// TIA Portal project "SSA-3GHz_V18" (V18) (continued)
REGION Network 10: PS_OK
   RUNG wire#powerrail
      Contact( "DigitalInputs".PS_OK.DigitalIN.NegLogic )
      I_Contact( "DigitalInputs".PS_OK.DigitalIN.PhysIn )
      wire#w1
      Coil( "DigitalInputs".PS_OK.DigitalIN.Out )
   END_RUNG
   RUNG wire#powerrail
      I_Contact( "DigitalInputs".PS_OK.DigitalIN.NegLogic )
      Contact( "DigitalInputs".PS_OK.DigitalIN.PhysIn )
   END_RUNG wire#w1
   // the same network as SCL:
   "DigitalInputs".PS_OK.DigitalIN.Out := ("DigitalInputs".PS_OK.DigitalIN.NegLogic AND NOT "DigitalInputs".PS_OK.DigitalIN.PhysIn) OR (NOT "DigitalInputs".PS_OK.DigitalIN.NegLogic AND "DigitalInputs".PS_OK.DigitalIN.PhysIn);
END_REGION

REGION Network 11: CoolingWtrOK
   RUNG wire#powerrail
      Contact( "CoolingWtrOK" )
      Coil( "DigitalInputs".CoolingWtrOK.DigitalIN.PhysIn )
   END_RUNG
   // the same network as SCL:
   "DigitalInputs".CoolingWtrOK.DigitalIN.PhysIn := "CoolingWtrOK";
END_REGION

REGION Network 12: CoolingWtrOK
   RUNG wire#powerrail
      Contact( "DigitalInputs".CoolingWtrOK.DigitalIN.NegLogic )
      I_Contact( "DigitalInputs".CoolingWtrOK.DigitalIN.PhysIn )
      wire#w1
      Coil( "DigitalInputs".CoolingWtrOK.DigitalIN.Out )
   END_RUNG
   RUNG wire#powerrail
      I_Contact( "DigitalInputs".CoolingWtrOK.DigitalIN.NegLogic )
      Contact( "DigitalInputs".CoolingWtrOK.DigitalIN.PhysIn )
   END_RUNG wire#w1
   // the same network as SCL:
   "DigitalInputs".CoolingWtrOK.DigitalIN.Out := ("DigitalInputs".CoolingWtrOK.DigitalIN.NegLogic AND NOT "DigitalInputs".CoolingWtrOK.DigitalIN.PhysIn) OR (NOT "DigitalInputs".CoolingWtrOK.DigitalIN.NegLogic AND "DigitalInputs".CoolingWtrOK.DigitalIN.PhysIn);
END_REGION

REGION Network 13: FanOK
   RUNG wire#powerrail
      Contact( "FanOK" )
      Coil( "DigitalInputs".FanOK.DigitalIN.PhysIn )
   END_RUNG
   // the same network as SCL:
   "DigitalInputs".FanOK.DigitalIN.PhysIn := "FanOK";
END_REGION

REGION Network 14: FanOK
   RUNG wire#powerrail
      Contact( "DigitalInputs".FanOK.DigitalIN.NegLogic )
      I_Contact( "DigitalInputs".FanOK.DigitalIN.PhysIn )
      wire#w1
      Coil( "DigitalInputs".FanOK.DigitalIN.Out )
   END_RUNG
   RUNG wire#powerrail
      I_Contact( "DigitalInputs".FanOK.DigitalIN.NegLogic )
      Contact( "DigitalInputs".FanOK.DigitalIN.PhysIn )
   END_RUNG wire#w1
   // the same network as SCL:
   "DigitalInputs".FanOK.DigitalIN.Out := ("DigitalInputs".FanOK.DigitalIN.NegLogic AND NOT "DigitalInputs".FanOK.DigitalIN.PhysIn) OR (NOT "DigitalInputs".FanOK.DigitalIN.NegLogic AND "DigitalInputs".FanOK.DigitalIN.PhysIn);
END_REGION

REGION Network 15: ExtIntlkOK
   RUNG wire#powerrail
      Contact( "ExtIntlkOK" )
      Coil( "DigitalInputs".ExtIntlkOK.DigitalIN.PhysIn )
   END_RUNG
   // the same network as SCL:
   "DigitalInputs".ExtIntlkOK.DigitalIN.PhysIn := "ExtIntlkOK";
END_REGION

REGION Network 16: ExtIntlkOK
   RUNG wire#powerrail
      Contact( "DigitalInputs".ExtIntlkOK.DigitalIN.NegLogic )
      I_Contact( "DigitalInputs".ExtIntlkOK.DigitalIN.PhysIn )
      wire#w1
      Coil( "DigitalInputs".ExtIntlkOK.DigitalIN.Out )
   END_RUNG
   RUNG wire#powerrail
      I_Contact( "DigitalInputs".ExtIntlkOK.DigitalIN.NegLogic )
      Contact( "DigitalInputs".ExtIntlkOK.DigitalIN.PhysIn )
   END_RUNG wire#w1
   // the same network as SCL:
   "DigitalInputs".ExtIntlkOK.DigitalIN.Out := ("DigitalInputs".ExtIntlkOK.DigitalIN.NegLogic AND NOT "DigitalInputs".ExtIntlkOK.DigitalIN.PhysIn) OR (NOT "DigitalInputs".ExtIntlkOK.DigitalIN.NegLogic AND "DigitalInputs".ExtIntlkOK.DigitalIN.PhysIn);
END_REGION
END_FUNCTION

FUNCTION "ProcessAI" : Void   // FC401, LAD
{ S7_Optimized_Access := 'TRUE' }
VERSION : 0.1
   VAR_TEMP
      tmpR : Real;
   END_VAR
BEGIN

REGION Network 1: U drain_RBK
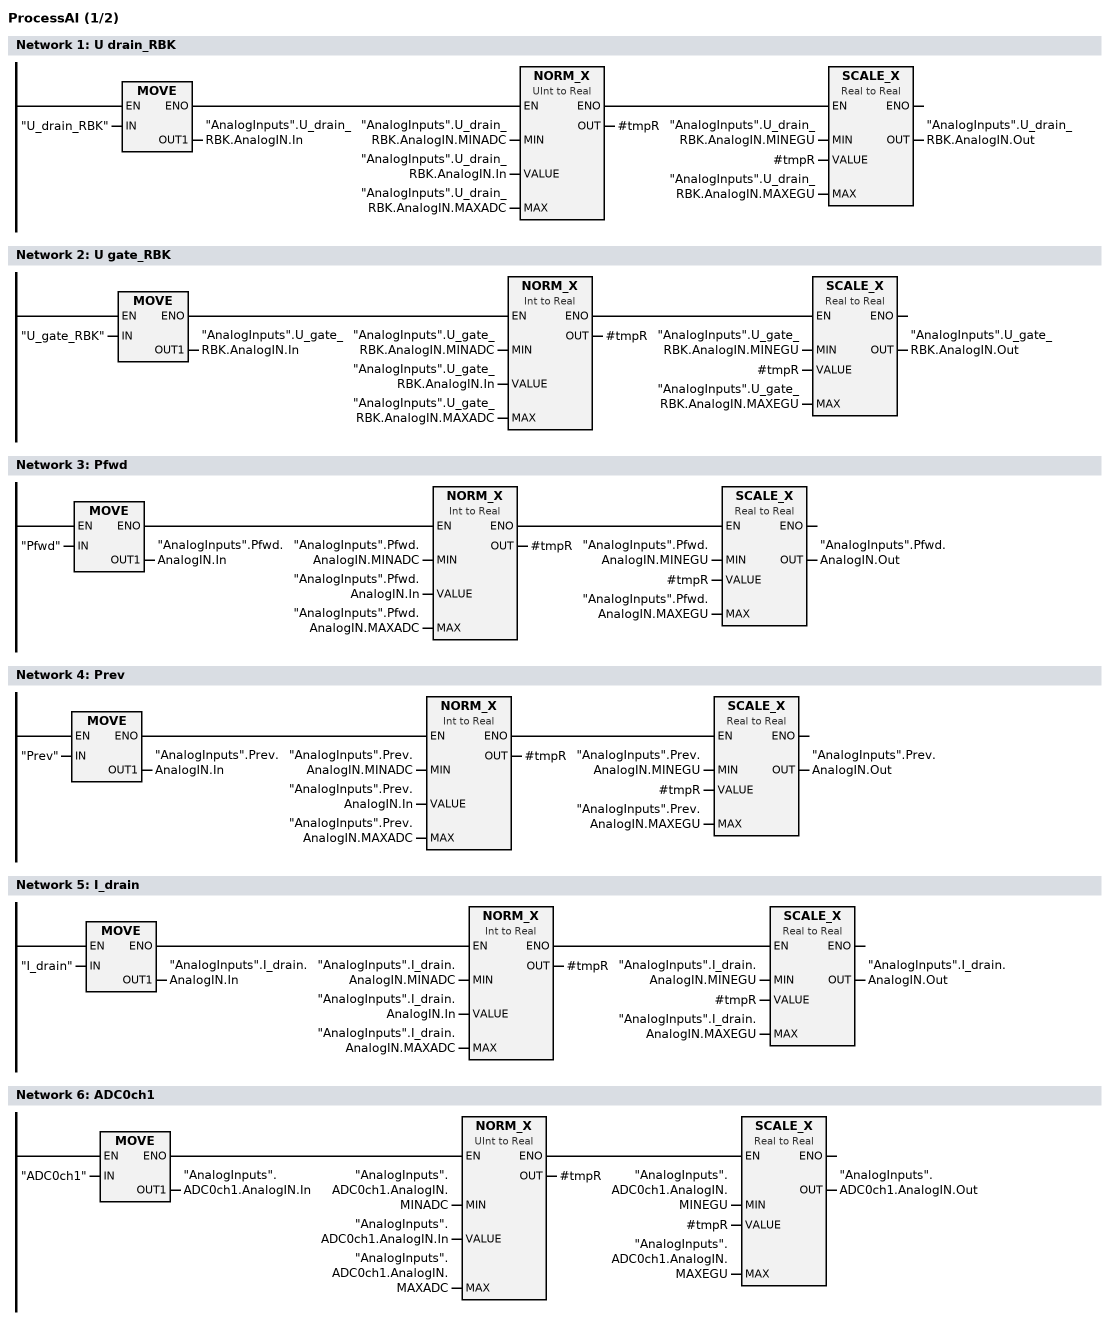
   RUNG wire#powerrail
      Move(in := "U_drain_RBK", out1 => "AnalogInputs".U_drain_RBK.AnalogIN.In)
      { S7_Templates := "[SrcType := UInt, DestType := Real]" } Normalize(min := "AnalogInputs".U_drain_RBK.AnalogIN.MINADC, value := "AnalogInputs".U_drain_RBK.AnalogIN.In, max := "AnalogInputs".U_drain_RBK.AnalogIN.MAXADC, out => #tmpR)
      { S7_Templates := "[SrcType := Real, DestType := Real]" } Scale(min := "AnalogInputs".U_drain_RBK.AnalogIN.MINEGU, value := #tmpR, max := "AnalogInputs".U_drain_RBK.AnalogIN.MAXEGU, out => "AnalogInputs".U_drain_RBK.AnalogIN.Out)
   END_RUNG
   // the same network as SCL:
   "AnalogInputs".U_drain_RBK.AnalogIN.In := "U_drain_RBK";
   #tmpR := NORM_X(MIN := "AnalogInputs".U_drain_RBK.AnalogIN.MINADC, VALUE := "AnalogInputs".U_drain_RBK.AnalogIN.In, MAX := "AnalogInputs".U_drain_RBK.AnalogIN.MAXADC);
   "AnalogInputs".U_drain_RBK.AnalogIN.Out := SCALE_X(MIN := "AnalogInputs".U_drain_RBK.AnalogIN.MINEGU, VALUE := #tmpR, MAX := "AnalogInputs".U_drain_RBK.AnalogIN.MAXEGU);
END_REGION

REGION Network 2: U gate_RBK
   RUNG wire#powerrail
      Move(in := "U_gate_RBK", out1 => "AnalogInputs".U_gate_RBK.AnalogIN.In)
      { S7_Templates := "[SrcType := Int, DestType := Real]" } Normalize(min := "AnalogInputs".U_gate_RBK.AnalogIN.MINADC, value := "AnalogInputs".U_gate_RBK.AnalogIN.In, max := "AnalogInputs".U_gate_RBK.AnalogIN.MAXADC, out => #tmpR)
      { S7_Templates := "[SrcType := Real, DestType := Real]" } Scale(min := "AnalogInputs".U_gate_RBK.AnalogIN.MINEGU, value := #tmpR, max := "AnalogInputs".U_gate_RBK.AnalogIN.MAXEGU, out => "AnalogInputs".U_gate_RBK.AnalogIN.Out)
   END_RUNG
   // the same network as SCL:
   "AnalogInputs".U_gate_RBK.AnalogIN.In := "U_gate_RBK";
   #tmpR := NORM_X(MIN := "AnalogInputs".U_gate_RBK.AnalogIN.MINADC, VALUE := "AnalogInputs".U_gate_RBK.AnalogIN.In, MAX := "AnalogInputs".U_gate_RBK.AnalogIN.MAXADC);
   "AnalogInputs".U_gate_RBK.AnalogIN.Out := SCALE_X(MIN := "AnalogInputs".U_gate_RBK.AnalogIN.MINEGU, VALUE := #tmpR, MAX := "AnalogInputs".U_gate_RBK.AnalogIN.MAXEGU);
END_REGION

REGION Network 3: Pfwd
   RUNG wire#powerrail
      Move(in := "Pfwd", out1 => "AnalogInputs".Pfwd.AnalogIN.In)
      { S7_Templates := "[SrcType := Int, DestType := Real]" } Normalize(min := "AnalogInputs".Pfwd.AnalogIN.MINADC, value := "AnalogInputs".Pfwd.AnalogIN.In, max := "AnalogInputs".Pfwd.AnalogIN.MAXADC, out => #tmpR)
      { S7_Templates := "[SrcType := Real, DestType := Real]" } Scale(min := "AnalogInputs".Pfwd.AnalogIN.MINEGU, value := #tmpR, max := "AnalogInputs".Pfwd.AnalogIN.MAXEGU, out => "AnalogInputs".Pfwd.AnalogIN.Out)
   END_RUNG
   // the same network as SCL:
   "AnalogInputs".Pfwd.AnalogIN.In := "Pfwd";
   #tmpR := NORM_X(MIN := "AnalogInputs".Pfwd.AnalogIN.MINADC, VALUE := "AnalogInputs".Pfwd.AnalogIN.In, MAX := "AnalogInputs".Pfwd.AnalogIN.MAXADC);
   "AnalogInputs".Pfwd.AnalogIN.Out := SCALE_X(MIN := "AnalogInputs".Pfwd.AnalogIN.MINEGU, VALUE := #tmpR, MAX := "AnalogInputs".Pfwd.AnalogIN.MAXEGU);
END_REGION

REGION Network 4: Prev
   RUNG wire#powerrail
      Move(in := "Prev", out1 => "AnalogInputs".Prev.AnalogIN.In)
      { S7_Templates := "[SrcType := Int, DestType := Real]" } Normalize(min := "AnalogInputs".Prev.AnalogIN.MINADC, value := "AnalogInputs".Prev.AnalogIN.In, max := "AnalogInputs".Prev.AnalogIN.MAXADC, out => #tmpR)
      { S7_Templates := "[SrcType := Real, DestType := Real]" } Scale(min := "AnalogInputs".Prev.AnalogIN.MINEGU, value := #tmpR, max := "AnalogInputs".Prev.AnalogIN.MAXEGU, out => "AnalogInputs".Prev.AnalogIN.Out)
   END_RUNG
   // the same network as SCL:
   "AnalogInputs".Prev.AnalogIN.In := "Prev";
   #tmpR := NORM_X(MIN := "AnalogInputs".Prev.AnalogIN.MINADC, VALUE := "AnalogInputs".Prev.AnalogIN.In, MAX := "AnalogInputs".Prev.AnalogIN.MAXADC);
   "AnalogInputs".Prev.AnalogIN.Out := SCALE_X(MIN := "AnalogInputs".Prev.AnalogIN.MINEGU, VALUE := #tmpR, MAX := "AnalogInputs".Prev.AnalogIN.MAXEGU);
END_REGION

REGION Network 5: I_drain
   RUNG wire#powerrail
      Move(in := "I_drain", out1 => "AnalogInputs".I_drain.AnalogIN.In)
      { S7_Templates := "[SrcType := Int, DestType := Real]" } Normalize(min := "AnalogInputs".I_drain.AnalogIN.MINADC, value := "AnalogInputs".I_drain.AnalogIN.In, max := "AnalogInputs".I_drain.AnalogIN.MAXADC, out => #tmpR)
      { S7_Templates := "[SrcType := Real, DestType := Real]" } Scale(min := "AnalogInputs".I_drain.AnalogIN.MINEGU, value := #tmpR, max := "AnalogInputs".I_drain.AnalogIN.MAXEGU, out => "AnalogInputs".I_drain.AnalogIN.Out)
   END_RUNG
   // the same network as SCL:
   "AnalogInputs".I_drain.AnalogIN.In := "I_drain";
   #tmpR := NORM_X(MIN := "AnalogInputs".I_drain.AnalogIN.MINADC, VALUE := "AnalogInputs".I_drain.AnalogIN.In, MAX := "AnalogInputs".I_drain.AnalogIN.MAXADC);
   "AnalogInputs".I_drain.AnalogIN.Out := SCALE_X(MIN := "AnalogInputs".I_drain.AnalogIN.MINEGU, VALUE := #tmpR, MAX := "AnalogInputs".I_drain.AnalogIN.MAXEGU);
END_REGION

REGION Network 6: ADC0ch1
   RUNG wire#powerrail
      Move(in := "ADC0ch1", out1 => "AnalogInputs".ADC0ch1.AnalogIN.In)
      { S7_Templates := "[SrcType := UInt, DestType := Real]" } Normalize(min := "AnalogInputs".ADC0ch1.AnalogIN.MINADC, value := "AnalogInputs".ADC0ch1.AnalogIN.In, max := "AnalogInputs".ADC0ch1.AnalogIN.MAXADC, out => #tmpR)
      { S7_Templates := "[SrcType := Real, DestType := Real]" } Scale(min := "AnalogInputs".ADC0ch1.AnalogIN.MINEGU, value := #tmpR, max := "AnalogInputs".ADC0ch1.AnalogIN.MAXEGU, out => "AnalogInputs".ADC0ch1.AnalogIN.Out)
   END_RUNG
   // the same network as SCL:
   "AnalogInputs".ADC0ch1.AnalogIN.In := "ADC0ch1";
   #tmpR := NORM_X(MIN := "AnalogInputs".ADC0ch1.AnalogIN.MINADC, VALUE := "AnalogInputs".ADC0ch1.AnalogIN.In, MAX := "AnalogInputs".ADC0ch1.AnalogIN.MAXADC);
   "AnalogInputs".ADC0ch1.AnalogIN.Out := SCALE_X(MIN := "AnalogInputs".ADC0ch1.AnalogIN.MINEGU, VALUE := #tmpR, MAX := "AnalogInputs".ADC0ch1.AnalogIN.MAXEGU);
END_REGION

REGION Network 7: Pfwd in dBm
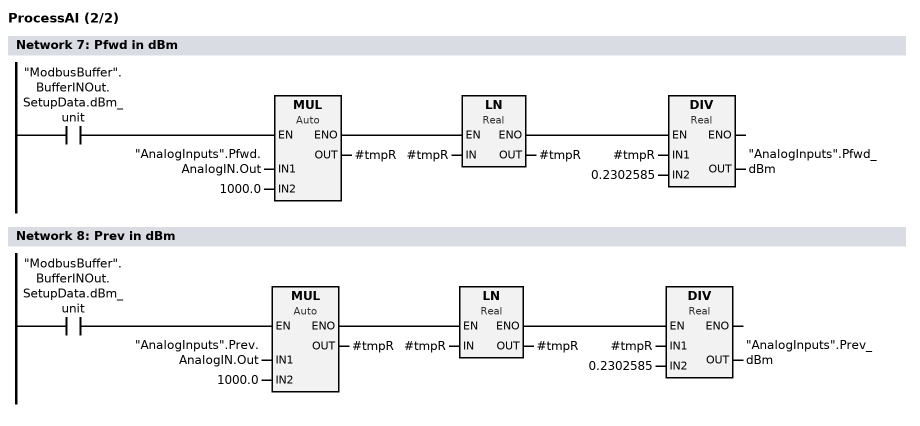
   IF "ModbusBuffer".BufferINOut.SetupData.dBm_unit THEN
       #tmpR := "AnalogInputs".Pfwd.AnalogIN.Out * 1000.0;
       #tmpR := LN(#tmpR);
       "AnalogInputs".Pfwd_dBm := #tmpR / 0.2302585;
   END_IF;
END_REGION

REGION Network 8: Prev in dBm
   IF "ModbusBuffer".BufferINOut.SetupData.dBm_unit THEN
       #tmpR := "AnalogInputs".Prev.AnalogIN.Out * 1000.0;
       #tmpR := LN(#tmpR);
       "AnalogInputs".Prev_dBm := #tmpR / 0.2302585;
   END_IF;
END_REGION
END_FUNCTION

FUNCTION "ProcessAO" : Void   // FC402, LAD
{ S7_Optimized_Access := 'TRUE' }
VERSION : 0.1
   VAR_TEMP
      tmpR : Real;
   END_VAR
BEGIN

REGION Network 1: U drain
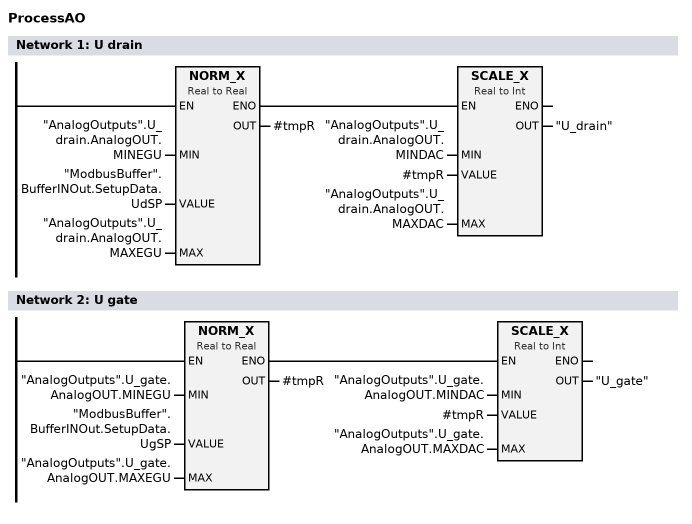
   RUNG wire#powerrail
      { S7_Templates := "[SrcType := Real, DestType := Real]" } Normalize(min := "AnalogOutputs".U_drain.AnalogOUT.MINEGU, value := "ModbusBuffer".BufferINOut.SetupData.UdSP, max := "AnalogOutputs".U_drain.AnalogOUT.MAXEGU, out => #tmpR)
      { S7_Templates := "[SrcType := Real, DestType := Int]" } Scale(min := "AnalogOutputs".U_drain.AnalogOUT.MINDAC, value := #tmpR, max := "AnalogOutputs".U_drain.AnalogOUT.MAXDAC, out => "U_drain")
   END_RUNG
   // the same network as SCL:
   #tmpR := NORM_X(MIN := "AnalogOutputs".U_drain.AnalogOUT.MINEGU, VALUE := "ModbusBuffer".BufferINOut.SetupData.UdSP, MAX := "AnalogOutputs".U_drain.AnalogOUT.MAXEGU);
   "U_drain" := SCALE_X(MIN := "AnalogOutputs".U_drain.AnalogOUT.MINDAC, VALUE := #tmpR, MAX := "AnalogOutputs".U_drain.AnalogOUT.MAXDAC);
END_REGION

REGION Network 2: U gate
   RUNG wire#powerrail
      { S7_Templates := "[SrcType := Real, DestType := Real]" } Normalize(min := "AnalogOutputs".U_gate.AnalogOUT.MINEGU, value := "ModbusBuffer".BufferINOut.SetupData.UgSP, max := "AnalogOutputs".U_gate.AnalogOUT.MAXEGU, out => #tmpR)
      { S7_Templates := "[SrcType := Real, DestType := Int]" } Scale(min := "AnalogOutputs".U_gate.AnalogOUT.MINDAC, value := #tmpR, max := "AnalogOutputs".U_gate.AnalogOUT.MAXDAC, out => "U_gate")
   END_RUNG
   // the same network as SCL:
   #tmpR := NORM_X(MIN := "AnalogOutputs".U_gate.AnalogOUT.MINEGU, VALUE := "ModbusBuffer".BufferINOut.SetupData.UgSP, MAX := "AnalogOutputs".U_gate.AnalogOUT.MAXEGU);
   "U_gate" := SCALE_X(MIN := "AnalogOutputs".U_gate.AnalogOUT.MINDAC, VALUE := #tmpR, MAX := "AnalogOutputs".U_gate.AnalogOUT.MAXDAC);
END_REGION
END_FUNCTION

FUNCTION "ProcessDO" : Void   // FC450, LAD
{ S7_Optimized_Access := 'TRUE' }
VERSION : 0.1
BEGIN

REGION Network 1: RF switcch
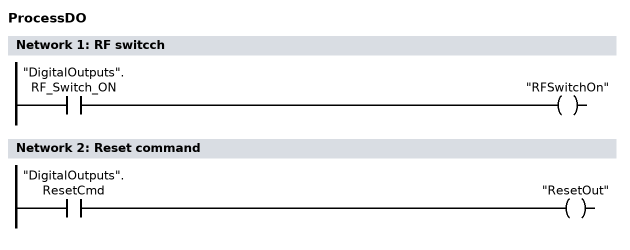
   RUNG wire#powerrail
      Contact( "DigitalOutputs".RF_Switch_ON )
      Coil( "RFSwitchOn" )
   END_RUNG
   // the same network as SCL:
   "RFSwitchOn" := "DigitalOutputs".RF_Switch_ON;
END_REGION

REGION Network 2: Reset command
   RUNG wire#powerrail
      Contact( "DigitalOutputs".ResetCmd )
      Coil( "ResetOut" )
   END_RUNG
   // the same network as SCL:
   "ResetOut" := "DigitalOutputs".ResetCmd;
END_REGION
END_FUNCTION

FUNCTION "CalcTransistorV" : Void   // FC500, SCL
{ S7_Optimized_Access := 'TRUE' }
VERSION : 0.1
   VAR_INPUT
      NominalPwr : Real;
      size : Int;   // max size if the lookup table. Valid data until Pwr != 0
   END_VAR
   VAR_OUTPUT
      UdSP : Real;
      UgSP : Real;
   END_VAR
   VAR_TEMP
      Pwr : Real;
      Ud : Real;
      Ug : Real;
      K : Real;
      i : Int;
   END_VAR
BEGIN
   (*
   Calculate the Darin and gate voltages based on the nominal power
   *)
   IF "ModbusBuffer".BufferINOut.SetupData.dBm_unit THEN
       "ModbusBuffer".BufferINOut.SetupData.NominalPower := EXP("ModbusBuffer".BufferINOut.SetupData.NominalPower_dBm* 0.2302585) / 1000.0;
   ELSE
       "ModbusBuffer".BufferINOut.SetupData.NominalPower_dBm := 10.0 * LN(1000.0 *"ModbusBuffer".BufferINOut.SetupData.NominalPower)/ 2.302585;
   END_IF;

   IF #NominalPwr <= "ModbusBuffer".BufferINOut.LookupTable.Pwr[0] THEN
       #UdSP := "ModbusBuffer".BufferINOut.LookupTable.Ud[0];
       #UgSP := "ModbusBuffer".BufferINOut.LookupTable.Ug[0];
   ELSE
       FOR #i := 1 TO #size-1 DO
       // Statement section FOR
           #Pwr := "ModbusBuffer".BufferINOut.LookupTable.Pwr[#i];
           IF #Pwr = 0 THEN
               //the end of table marker
               #UdSP := "ModbusBuffer".BufferINOut.LookupTable.Ud[#i - 1];
               #UgSP := "ModbusBuffer".BufferINOut.LookupTable.Ug[#i - 1];
               RETURN;
           END_IF;
           IF #NominalPwr > #Pwr THEN
               CONTINUE;
           END_IF;
           #K := (#NominalPwr - "ModbusBuffer".BufferINOut.LookupTable.Pwr[#i - 1]) / (#Pwr - "ModbusBuffer".BufferINOut.LookupTable.Pwr[#i - 1]);
           #UdSP := "ModbusBuffer".BufferINOut.LookupTable.Ud[#i-1] + #K * ("ModbusBuffer".BufferINOut.LookupTable.Ud[#i] - "ModbusBuffer".BufferINOut.LookupTable.Ud[#i-1]);
           #UgSP := "ModbusBuffer".BufferINOut.LookupTable.Ug[#i - 1] + #K * ("ModbusBuffer".BufferINOut.LookupTable.Ug[#i] - "ModbusBuffer".BufferINOut.LookupTable.Ug[#i - 1]);
           RETURN;
       END_FOR;
       #UdSP := "ModbusBuffer".BufferINOut.LookupTable.Ud[#size-1];
       #UgSP := "ModbusBuffer".BufferINOut.LookupTable.Ug[#size-1];
   END_IF;
END_FUNCTION

FUNCTION "Interlocks" : Void   // FC600, LAD
{ S7_Optimized_Access := 'TRUE' }
VERSION : 0.1
BEGIN

REGION Network 1: RF Switch
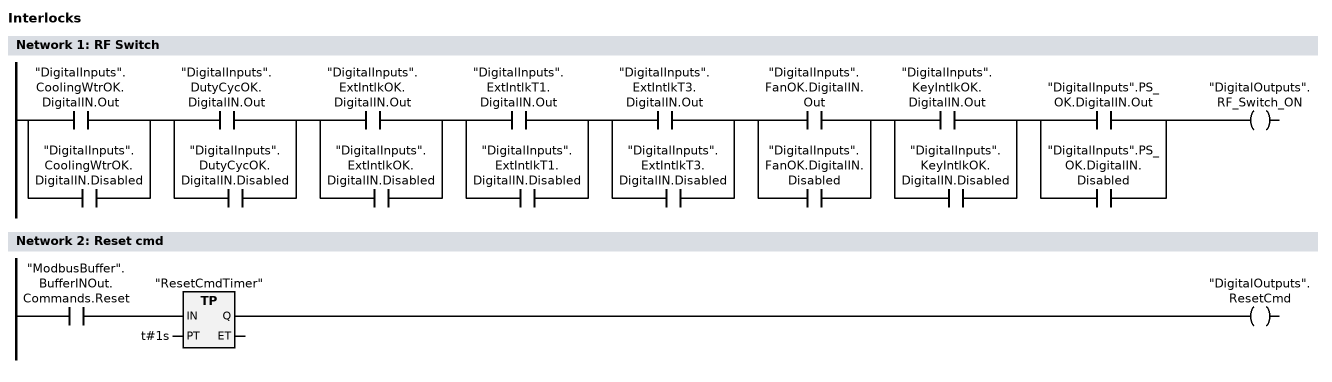
   RUNG wire#powerrail
      Contact( "DigitalInputs".CoolingWtrOK.DigitalIN.Out )
      wire#w1
      Contact( "DigitalInputs".DutyCycOK.DigitalIN.Out )
      wire#w2
      Contact( "DigitalInputs".ExtIntlkOK.DigitalIN.Out )
      wire#w3
      Contact( "DigitalInputs".ExtIntlkT1.DigitalIN.Out )
      wire#w4
      Contact( "DigitalInputs".ExtIntlkT3.DigitalIN.Out )
      wire#w5
      Contact( "DigitalInputs".FanOK.DigitalIN.Out )
      wire#w6
      Contact( "DigitalInputs".KeyIntlkOK.DigitalIN.Out )
      wire#w7
      Contact( "DigitalInputs".PS_OK.DigitalIN.Out )
      wire#w8
      Coil( "DigitalOutputs".RF_Switch_ON )
   END_RUNG
   RUNG wire#powerrail
      Contact( "DigitalInputs".CoolingWtrOK.DigitalIN.Disabled )
   END_RUNG wire#w1
   RUNG wire#w1
      Contact( "DigitalInputs".DutyCycOK.DigitalIN.Disabled )
   END_RUNG wire#w2
   RUNG wire#w2
      Contact( "DigitalInputs".ExtIntlkOK.DigitalIN.Disabled )
   END_RUNG wire#w3
   RUNG wire#w3
      Contact( "DigitalInputs".ExtIntlkT1.DigitalIN.Disabled )
   END_RUNG wire#w4
   RUNG wire#w4
      Contact( "DigitalInputs".ExtIntlkT3.DigitalIN.Disabled )
   END_RUNG wire#w5
   RUNG wire#w5
      Contact( "DigitalInputs".FanOK.DigitalIN.Disabled )
   END_RUNG wire#w6
   RUNG wire#w6
      Contact( "DigitalInputs".KeyIntlkOK.DigitalIN.Disabled )
   END_RUNG wire#w7
   RUNG wire#w7
      Contact( "DigitalInputs".PS_OK.DigitalIN.Disabled )
   END_RUNG wire#w8
   // the same network as SCL:
   "DigitalOutputs".RF_Switch_ON := ("DigitalInputs".CoolingWtrOK.DigitalIN.Out OR "DigitalInputs".CoolingWtrOK.DigitalIN.Disabled) AND ("DigitalInputs".DutyCycOK.DigitalIN.Out OR "DigitalInputs".DutyCycOK.DigitalIN.Disabled) AND ("DigitalInputs".ExtIntlkOK.DigitalIN.Out OR "DigitalInputs".ExtIntlkOK.DigitalIN.Disabled) AND ("DigitalInputs".ExtIntlkT1.DigitalIN.Out OR "DigitalInputs".ExtIntlkT1.DigitalIN.Disabled) AND ("DigitalInputs".ExtIntlkT3.DigitalIN.Out OR "DigitalInputs".ExtIntlkT3.DigitalIN.Disabled) AND ("DigitalInputs".FanOK.DigitalIN.Out OR "DigitalInputs".FanOK.DigitalIN.Disabled) AND ("DigitalInputs".KeyIntlkOK.DigitalIN.Out OR "DigitalInputs".KeyIntlkOK.DigitalIN.Disabled) AND ("DigitalInputs".PS_OK.DigitalIN.Out OR "DigitalInputs".PS_OK.DigitalIN.Disabled);
END_REGION

REGION Network 2: Reset cmd
   "ResetCmdTimer".TP(IN := "ModbusBuffer".BufferINOut.Commands.Reset, PT := t#1s);
   "DigitalOutputs".ResetCmd := "ResetCmdTimer".Q;
END_REGION
END_FUNCTION

ORGANIZATION_BLOCK "Main"   // OB1, LAD, ProgramCycle
TITLE = "Main Program Sweep (Cycle)"
{ S7_Optimized_Access := 'TRUE' }
VERSION : 0.1
   VAR_INPUT
      Initial_Call : Bool;   // Initial call of this OB
      Remanence : Bool;   // =True, if remanent data are available
   END_VAR
BEGIN

REGION Network 1: Setup
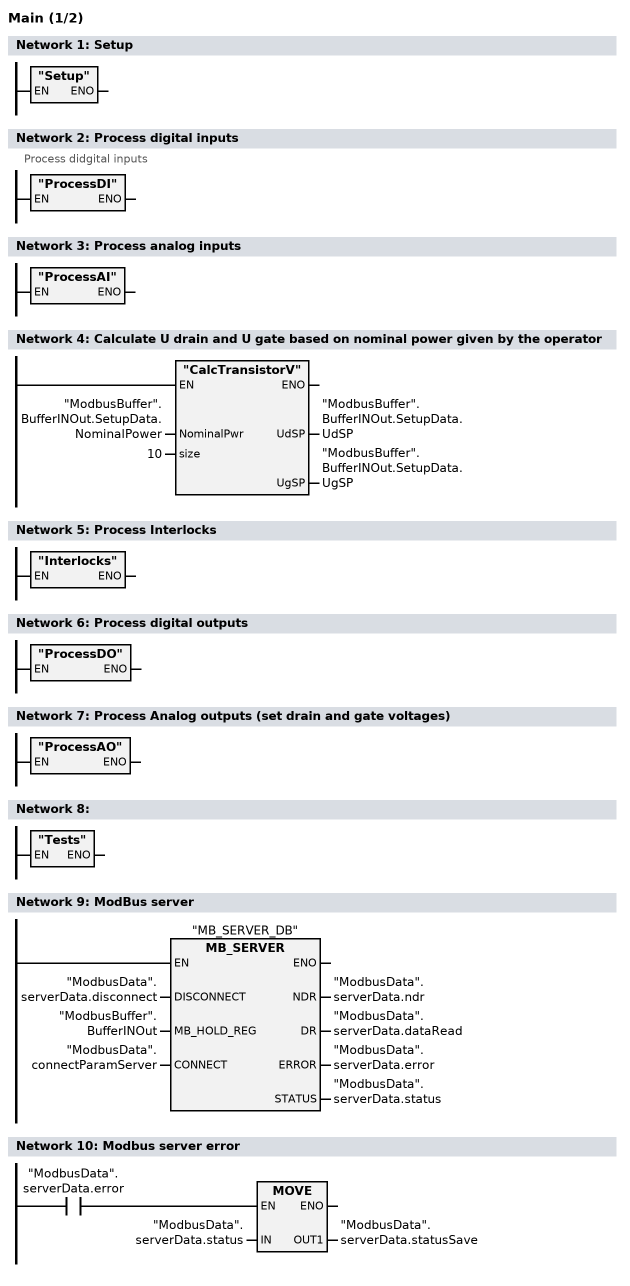
   RUNG wire#powerrail
      "Setup"()
   END_RUNG
   // the same network as SCL:
   "Setup"();
END_REGION

REGION Network 2: Process digital inputs
   // Process didgital inputs
   RUNG wire#powerrail
      "ProcessDI"()
   END_RUNG
   // the same network as SCL:
   "ProcessDI"();
END_REGION

REGION Network 3: Process analog inputs
   RUNG wire#powerrail
      "ProcessAI"()
   END_RUNG
   // the same network as SCL:
   "ProcessAI"();
END_REGION

REGION Network 4: Calculate U drain and U gate based on nominal power given by the operator
   RUNG wire#powerrail
      "CalcTransistorV"(NominalPwr := "ModbusBuffer".BufferINOut.SetupData.NominalPower, size := 10, UdSP => "ModbusBuffer".BufferINOut.SetupData.UdSP, UgSP => "ModbusBuffer".BufferINOut.SetupData.UgSP)
   END_RUNG
   // the same network as SCL:
   "CalcTransistorV"(NominalPwr := "ModbusBuffer".BufferINOut.SetupData.NominalPower,
                     size := 10,
                     UdSP => "ModbusBuffer".BufferINOut.SetupData.UdSP,
                     UgSP => "ModbusBuffer".BufferINOut.SetupData.UgSP);
END_REGION

REGION Network 5: Process Interlocks
   RUNG wire#powerrail
      "Interlocks"()
   END_RUNG
   // the same network as SCL:
   "Interlocks"();
END_REGION

REGION Network 6: Process digital outputs
   RUNG wire#powerrail
      "ProcessDO"()
   END_RUNG
   // the same network as SCL:
   "ProcessDO"();
END_REGION

REGION Network 7: Process Analog outputs (set drain and gate voltages)
   RUNG wire#powerrail
      "ProcessAO"()
   END_RUNG
   // the same network as SCL:
   "ProcessAO"();
END_REGION

REGION Network 8
   RUNG wire#powerrail
      "Tests"()
   END_RUNG
   // the same network as SCL:
   "Tests"();
END_REGION

REGION Network 9: ModBus server
   "MB_SERVER_DB"(DISCONNECT := "ModbusData".serverData.disconnect,   // MB_SERVER
                  MB_HOLD_REG := "ModbusBuffer".BufferINOut,
                  CONNECT := "ModbusData".connectParamServer,
                  NDR => "ModbusData".serverData.ndr,
                  DR => "ModbusData".serverData.dataRead,
                  ERROR => "ModbusData".serverData.error,
                  STATUS => "ModbusData".serverData.status);
END_REGION

REGION Network 10: Modbus server error
   RUNG wire#powerrail
      Contact( "ModbusData".serverData.error )
      Move(in := "ModbusData".serverData.status, out1 => "ModbusData".serverData.statusSave)
   END_RUNG
   // the same network as SCL:
   IF "ModbusData".serverData.error THEN
       "ModbusData".serverData.statusSave := "ModbusData".serverData.status;
   END_IF;
END_REGION

REGION Network 11: Process data sent to the PLC via Modbus
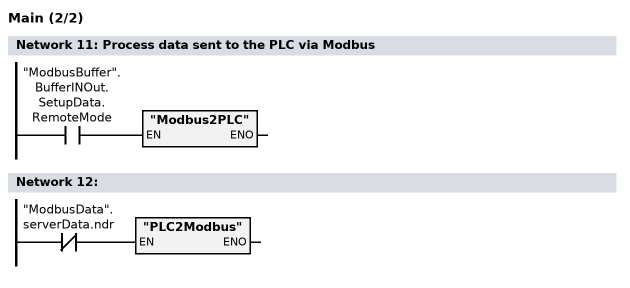
   RUNG wire#powerrail
      Contact( "ModbusBuffer".BufferINOut.SetupData.RemoteMode )
      "Modbus2PLC"()
   END_RUNG
   // the same network as SCL:
   IF "ModbusBuffer".BufferINOut.SetupData.RemoteMode THEN "Modbus2PLC"(); END_IF;
END_REGION

REGION Network 12
   RUNG wire#powerrail
      I_Contact( "ModbusData".serverData.ndr )
      "PLC2Modbus"()
   END_RUNG
   // the same network as SCL:
   IF NOT "ModbusData".serverData.ndr THEN "PLC2Modbus"(); END_IF;
END_REGION
END_ORGANIZATION_BLOCK

// folder: 5_T_CONFIG (S7-1200, S7-1500)

FUNCTION_BLOCK "SLI_FB_T_CONFIG"   // FB4, LAD
{ S7_Optimized_Access := 'TRUE' }
VERSION : 0.1
// Info: The example is meant to change the PROFINET  device name and IP address of the CPU via its PROFINET interface.
   VAR
      T_CONFIG_Instance : T_CONFIG;
      done : Bool;
      errorLocation : DWord;
   END_VAR
BEGIN

REGION Network 1: Set "start" to TRUE to configure the PROFINET interface.
   // NOTE! Before using the example:
   // 
   // Condition:
   // 1) Open the device view of the CPU "> Properties > PROFINET interface > Ethernet addresses > PROFINET". 
   // 2) To set the device name: Activate the following options: 
   // - "IP address is set directly at the device". 
   // - "PROFINET device name is set directly at the device".
   // 
   // Regarding parameter INTERFACE ("hwid"):
   // - Change the value of "hwid" according to the identification number of the PROFINET interface of your local device (CPU). (Open "PLC tags > Show all tags > System constants. Look for a name like "<Local~PROFINET_interface_1>" with a Data type "Hw_Interface". The cell "value" contains the hwid.)
   // 
   // Info:
   // In the "header" (IF_CONF_HEADER):
   // - SubfieldCount = 2: Indicates that two additional structures ("deviceIP" and "deviceName") are used below.
   // 
   // In the structure "deviceIP" (system data type IF_CONF_v4):
   // - Lenght = 18: Information on overall length of the structure (12 bytes for the device IP + 6 bytes for the parameters Id, Length and Mode)
   // - Mode = 1: Permanent change of the device IP.
   // - InterfaceAddress, SubnetMask, DefaultRouter: IP connection data.
   // 
   // In the structure "deviceName" (system data type IF_CONF_NOS):
   // - Lenght = 11: Information on overall length of the structure (5 bytes for the device name "myplc" + 6 bytes for the parameters Id, Length and Mode)
   // - Mode = 1: Permanent change of the device name in "myplc".
   // - NOS[1] ... NOS[5]: Device name (1 character / byte)
   // 
   // Note: Instead of an absolute length, you can use the default start value (Lenght = 0) for a dynamic length.
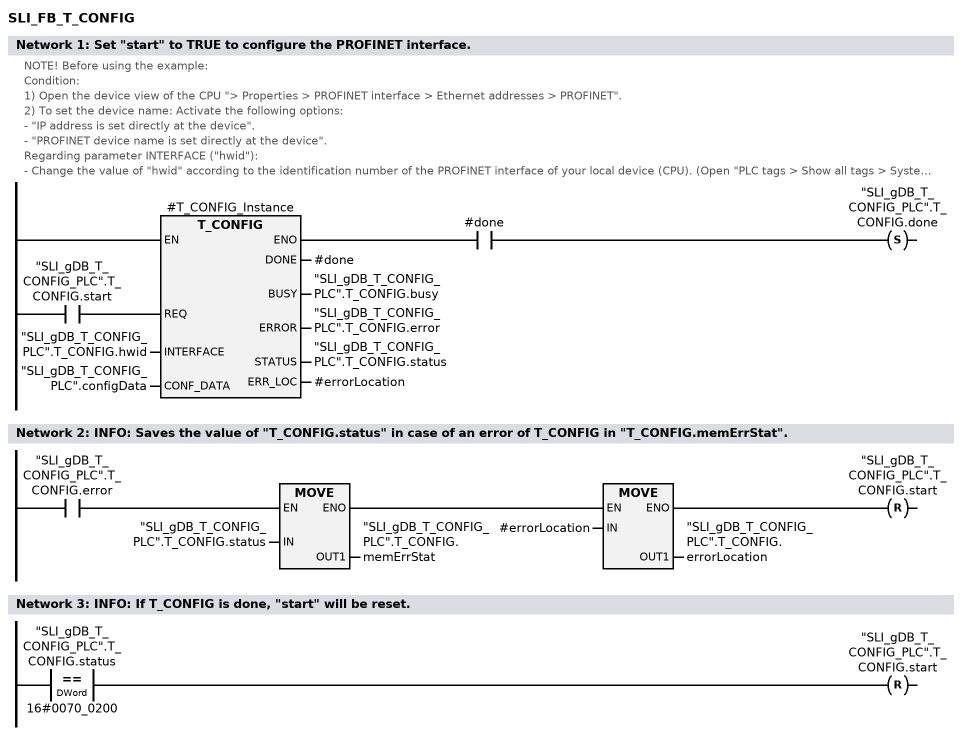
   // ENO of a box is taken as its EN; it also drops when the box reports an error
   #T_CONFIG_Instance(Req := "SLI_gDB_T_CONFIG_PLC".T_CONFIG.start,   // T_CONFIG
                      Interface := "SLI_gDB_T_CONFIG_PLC".T_CONFIG.hwid,
                      Conf_Data := "SLI_gDB_T_CONFIG_PLC".configData,
                      Done => #done,
                      Busy => "SLI_gDB_T_CONFIG_PLC".T_CONFIG.busy,
                      Error => "SLI_gDB_T_CONFIG_PLC".T_CONFIG.error,
                      Status => "SLI_gDB_T_CONFIG_PLC".T_CONFIG.status,
                      Err_Loc => #errorLocation);
   IF #done THEN "SLI_gDB_T_CONFIG_PLC".T_CONFIG.done := TRUE; END_IF;
END_REGION

REGION Network 2: INFO: Saves the value of "T_CONFIG.status" in case of an error of T_CONFIG in "T_CONFIG.memErrStat".
   RUNG wire#powerrail
      Contact( "SLI_gDB_T_CONFIG_PLC".T_CONFIG.error )
      Move(in := "SLI_gDB_T_CONFIG_PLC".T_CONFIG.status, out1 => "SLI_gDB_T_CONFIG_PLC".T_CONFIG.memErrStat)
      Move(in := #errorLocation, out1 => "SLI_gDB_T_CONFIG_PLC".T_CONFIG.errorLocation)
      R_Coil( "SLI_gDB_T_CONFIG_PLC".T_CONFIG.start )
   END_RUNG
   // the same network as SCL:
   IF "SLI_gDB_T_CONFIG_PLC".T_CONFIG.error THEN
       "SLI_gDB_T_CONFIG_PLC".T_CONFIG.memErrStat := "SLI_gDB_T_CONFIG_PLC".T_CONFIG.status;
       "SLI_gDB_T_CONFIG_PLC".T_CONFIG.errorLocation := #errorLocation;
       "SLI_gDB_T_CONFIG_PLC".T_CONFIG.start := FALSE;
   END_IF;
END_REGION

REGION Network 3: INFO: If T_CONFIG is done, "start" will be reset.
   RUNG wire#powerrail
      { S7_Templates := "SrcType := DWord" } EQ_Contact(in1 := "SLI_gDB_T_CONFIG_PLC".T_CONFIG.status, in2 := 16#0070_0200)
      R_Coil( "SLI_gDB_T_CONFIG_PLC".T_CONFIG.start )
   END_RUNG
   // the same network as SCL:
   IF "SLI_gDB_T_CONFIG_PLC".T_CONFIG.status = 16#0070_0200 THEN
       "SLI_gDB_T_CONFIG_PLC".T_CONFIG.start := FALSE;
   END_IF;
END_REGION
END_FUNCTION_BLOCK

(* ===== HMI "HMI_RT_1" =====
system functions are stored by id; their names below are inferred from use
connection "HMI_Connection_1": ETHERNET, SMART_S7_1200_OMS

HMI tags "Default tag table"
   "Tag_ScreenNumber" : UInt, internal
   "AnalogInputs_Pfwd_AnalogIN_Out" : Real = PLC AnalogInputs.Pfwd.AnalogIN.Out, 1 s
   "AnalogInputs_Prev_AnalogIN_Out" : Real = PLC AnalogInputs.Prev.AnalogIN.Out, 1 s
   "DigitalInputs_DutyCycOK_DigitalIN_Out" : Bool = PLC DigitalInputs.DutyCycOK.DigitalIN.Out, 1 s
   "DigitalInputs_KeyIntlkOK_DigitalIN_Out" : Bool = PLC DigitalInputs.KeyIntlkOK.DigitalIN.Out, 1 s
   "DigitalInputs_ExtIntlkT1_DigitalIN_Out" : Bool = PLC DigitalInputs.ExtIntlkT1.DigitalIN.Out, 1 s
   "DigitalInputs_ExtIntlkT3_DigitalIN_Out" : Bool = PLC DigitalInputs.ExtIntlkT3.DigitalIN.Out, 1 s
   "AnalogInputs_U_drain_RBK_AnalogIN_Out" : Real = PLC AnalogInputs.U_drain_RBK.AnalogIN.Out, 1 s
   "AnalogInputs_U_gate_RBK_AnalogIN_Out" : Real = PLC AnalogInputs.U_gate_RBK.AnalogIN.Out, 1 s
   "DigitalInputs_PS_OK_DigitalIN_Out" : Bool = PLC DigitalInputs.PS_OK.DigitalIN.Out, 1 s
   "DigitalInputs_CoolingWtrOK_DigitalIN_Out" : Bool = PLC DigitalInputs.CoolingWtrOK.DigitalIN.Out, 1 s
   "DigitalInputs_FanOK_DigitalIN_Out" : Bool = PLC DigitalInputs.FanOK.DigitalIN.Out, 1 s
   "DigitalInputs_ExtIntlkOK_DigitalIN_Out" : Bool = PLC DigitalInputs.ExtIntlkOK.DigitalIN.Out, 1 s
   "TestBlink" : Bool = PLC TestBlink AT %Q1.0, 1 s
   "AnalogInputs_U_gate_RBK_AnalogIN_VisuState" : Byte = PLC AnalogInputs.U_gate_RBK.AnalogIN.VisuState, 1 s
   "VisuTest" : Byte = PLC VisuTest AT %MB104, 1 s
   "DigitalInputs_DutyCycOK_DigitalIN_Disabled" : Bool = PLC DigitalInputs.DutyCycOK.DigitalIN.Disabled, 1 s
   "DigitalInputs_KeyIntlkOK_DigitalIN_Disabled" : Bool = PLC DigitalInputs.KeyIntlkOK.DigitalIN.Disabled, 1 s
   "DigitalInputs_ExtIntlkT1_DigitalIN_Disabled" : Bool = PLC DigitalInputs.ExtIntlkT1.DigitalIN.Disabled, 1 s
   "DigitalInputs_ExtIntlkT3_DigitalIN_Disabled" : Bool = PLC DigitalInputs.ExtIntlkT3.DigitalIN.Disabled, 1 s
   "DigitalInputs_PS_OK_DigitalIN_Disabled" : Bool = PLC DigitalInputs.PS_OK.DigitalIN.Disabled, 1 s
   "DigitalInputs_CoolingWtrOK_DigitalIN_Disabled" : Bool = PLC DigitalInputs.CoolingWtrOK.DigitalIN.Disabled, 1 s
   "DigitalInputs_FanOK_DigitalIN_Disabled" : Bool = PLC DigitalInputs.FanOK.DigitalIN.Disabled, 1 s
   "DigitalInputs_ExtIntlkOK_DigitalIN_Disabled" : Bool = PLC DigitalInputs.ExtIntlkOK.DigitalIN.Disabled, 1 s
   "ModbusBuffer_BufferINOut_SetupData_RemoteMode" : Bool = PLC ModbusBuffer.BufferINOut.SetupData.RemoteMode AT %DB101.DBX120.0, 1 s
   "ModbusBuffer_BufferINOut_SetupData_NominalPower" : Real = PLC ModbusBuffer.BufferINOut.SetupData.NominalPower AT %DB101.DBD122, 1 s
   "Counter_HMI" : UDInt = PLC Counter AT %MD100, 1 s

text list "Text_list_loc_rem": 0 'To Rem.'; 1 'To Loc.'

graphic list "Amplifier": 0 'Amplifier_grey_3'; 1 'Amplifier_blue_2'; 2 'Amplifier_green_2'; 3 'Amplifier_yellow_4'; 4 'Amplifier_red_3'

Template "Template" 480x272
   TextField "Template_Text field_1" at 94,6 size 23x37; Text 'P'
   TextField "Template_Text field_3" at 109,23 size 30x17; Text 'FWD'
   TextField "Template_Text field_5" at 258,8 size 23x37; Text 'P'
   TextField "Template_Text field_4" at 277,23 size 26x17; Text 'REV'
   Button "Alarms" at 1,46 size 63x44; TextOff 'Alarms'; PictureOff "AlarmDisplay_KTP400_Basic_PN_TR"; PictureOn "AlarmDisplay_KTP400_Basic_PN_TR"
      on Release: function_ef3f5d25("Alarm window_Unacknowledged", -1)
   Button "Template_Button_1" at 1,136 size 63x44; TextOff 'Text'
   Button "Template_Button_2" at 1,181 size 63x44; TextOff 'To Rem'; TextList "Text_list_loc_rem"
      on Release: InvertBit("ModbusBuffer_BufferINOut_SetupData_RemoteMode")
      ProcessValue <- "ModbusBuffer_BufferINOut_SetupData_RemoteMode"
   Button "Start screen" at 1,226 size 63x44; TextOff 'Start screen'; PictureOff "NavigateHome_KTP400_Basic_PN_TR"; PictureOn "NavigateHome_KTP400_Basic_PN_TR"
      on Release: ActivateScreen("Root screen", 0)
   DateTimeField "HmiScreenItemData" at 395,22 size 85x22
   DateTimeField "HmiScreenItemData_1" at 395,0 size 85x22
   GraphicView "Logo" at 0,0 size 94x45; Picture "Logo of HMI_1"
   Button "Template_Button_3" at 1,91 size 63x44; TextOff 'System'
      on Release: ActivateScreen("System screens", 0)
   TextField "Template_Text field_2" at 218,20 size 18x20; Text 'W'
   Group "Group" at 94,6 size 45x37
   Group "Group_1" at 258,8 size 45x37
   IOField "Template_I/O field_1" at 139,6 size 80x39; FormatPattern 9999
      ProcessValue <- "AnalogInputs_Pfwd_AnalogIN_Out"
   IOField "Template_I/O field_2" at 303,6 size 80x39; FormatPattern 9999
      ProcessValue <- "AnalogInputs_Prev_AnalogIN_Out"
   TextField "Template_Text field_6" at 382,20 size 18x20; Text 'W'

screen "Root screen" 480x272, template "Template"
   on GenerateScreen: SetTag("Tag_ScreenNumber", 1)
   TextField "Text field_1" at 69,239 size 70x20; Text 'Interlocks'
   TextField "Text field_2" at 146,229 size 75x20; Text 'Duty Cyc.'
      Appearance <- "DigitalInputs_DutyCycOK_DigitalIN_Out"
      Visibility <- "DigitalInputs_DutyCycOK_DigitalIN_Disabled"
   TextField "Text field_3" at 146,251 size 75x20; Text 'KeyIntlk'
      Appearance <- "DigitalInputs_KeyIntlkOK_DigitalIN_Out"
      Visibility <- "DigitalInputs_KeyIntlkOK_DigitalIN_Disabled"
   TextField "Text field_4" at 223,229 size 75x20; Text 'Intlk T1'
      Appearance <- "DigitalInputs_ExtIntlkT1_DigitalIN_Out"
      Visibility <- "DigitalInputs_ExtIntlkT1_DigitalIN_Disabled"
   TextField "Text field_5" at 223,251 size 75x20; Text 'Intlk T3'
      Appearance <- "DigitalInputs_ExtIntlkT3_DigitalIN_Out"
      Visibility <- "DigitalInputs_ExtIntlkT3_DigitalIN_Disabled"
   TextField "Text field_6" at 71,53 size 104x20; Text 'Nominal Power:'
   TextField "Text field_7" at 176,49 size 14x20; Text 'Text'
   IOField "I/O field_1" at 176,50 size 69x28; FormatPattern 9999
      ProcessValue <- "ModbusBuffer_BufferINOut_SetupData_NominalPower"
   Group "Group" at 69,82 size 19x20
   Group "Group_1" at 69,104 size 19x20
   IOField "I/O field_2" at 94,83 size 41x18; FormatPattern 99.9
      ProcessValue <- "AnalogInputs_U_drain_RBK_AnalogIN_Out"
   IOField "I/O field_3" at 94,105 size 41x18; FormatPattern 9.99
      ProcessValue <- "AnalogInputs_U_gate_RBK_AnalogIN_Out"
   TextField "Text field_13" at 300,229 size 75x20; Text 'PS_OK'
      Appearance <- "DigitalInputs_PS_OK_DigitalIN_Out"
      Visibility <- "DigitalInputs_PS_OK_DigitalIN_Disabled"
   TextField "Text field_14" at 300,251 size 75x20; Text 'CoolingWtr'
      Appearance <- "DigitalInputs_CoolingWtrOK_DigitalIN_Out"
      Visibility <- "DigitalInputs_CoolingWtrOK_DigitalIN_Disabled"
   TextField "Text field_15" at 377,229 size 75x20; Text 'Fan'
      Appearance <- "DigitalInputs_FanOK_DigitalIN_Out"
      Visibility <- "DigitalInputs_FanOK_DigitalIN_Disabled"
   TextField "Text field_16" at 377,251 size 75x20; Text 'ExtIntlk'
      Appearance <- "DigitalInputs_ExtIntlkOK_DigitalIN_Out"
      Visibility <- "DigitalInputs_ExtIntlkOK_DigitalIN_Disabled"
   TextField "Text field_17" at 75,143 size 37x20; Text 'RF In'
   TextField "Text field_18" at 408,145 size 47x20; Text 'RF Out'
   GraphicIOField "Graphic I/O field_2" at 197,91 size 175x128; PictureList "Amplifier"
      ProcessValue <- "VisuTest"
   Circle "Circle_1" at 421,71 size 31x31
      Appearance <- "TestBlink"
   IOField "I/O field_4" at 267,46 size 129x32; FormatPattern 9999999999
      ProcessValue <- "Counter_HMI"
   TextField "Text field_8" at 69,82 size 13x20; Text 'U'
   TextField "Text field_10" at 77,88 size 11x14; Text 'D'
   TextField "Text field_9" at 69,104 size 13x20; Text 'U'
   TextField "Text field_12" at 77,110 size 11x14; Text 'G'
   GraphicIOField "Graphic I/O field_1" at 141,143 size 45x23; PictureOff "JS Disconnecting Switch Off-RED"; PictureOn "JS Disconnecting Switch On-GREEN"
      ProcessValue <- "TestBlink"

screen "System screens" 480x272, template "Template"
   on GenerateScreen: SetTag("Tag_ScreenNumber", 2)
   TextField "HmiScreenItemData" at 106,145 size 332x22; Text 'System screens'
   Button "Back" at 65,46 size 136x30; TextOff 'Back'
      on Release: ActivateScreen("Root screen", 0)
   Button "SIMATIC PLC system diagnostics" at 65,77 size 136x30; TextOff 'SIMATIC PLC s...'
      on Release: ActivateScreen("SIMATIC PLC system diagnostics", 0)
   Button "Project information" at 65,108 size 136x30; TextOff 'Project informat...'
      on Release: ActivateScreen("Project information", 0)
   Button "System information" at 65,139 size 136x30; TextOff 'System informa...'
      on Release: ActivateScreen("System information", 0)

screen "SIMATIC PLC system diagnostics" 480x272, template "Template"
   on GenerateScreen: SetTag("Tag_ScreenNumber", 3)
   SysDiagControl "HmiScreenItemData" at 65,77 size 412x188
   Button "Back" at 65,46 size 136x30; TextOff 'Back'
      on Release: ActivateScreen("System screens", 0)

screen "Project information" 480x272, template "Template"
   on GenerateScreen: SetTag("Tag_ScreenNumber", 4)
   TextField "HmiScreenItemData" at 68,78 size 158x20; Text 'Project name:'
   TextField "HmiScreenItemData_1" at 230,78 size 246x20; Text 'SSA-3GHz'
   TextField "HmiScreenItemData_2" at 68,99 size 158x20; Text 'Created on:'
   TextField "HmiScreenItemData_3" at 230,99 size 246x20; Text '10/3/2022 1:09:17 PM'
   TextField "HmiScreenItemData_4" at 68,120 size 158x20; Text 'Author:'
   TextField "HmiScreenItemData_5" at 230,120 size 246x20; Text 'konrgaje'
   TextField "HmiScreenItemData_6" at 68,141 size 158x20; Text 'Description:'
   TextField "HmiScreenItemData_7" at 230,141 size 246x20; Text '(not configured)'
   Button "Back" at 65,46 size 136x30; TextOff 'Back'
      on Release: ActivateScreen("System screens", 0)

screen "System information" 480x272, template "Template"
   on GenerateScreen: SetTag("Tag_ScreenNumber", 5)
   TextField "HmiScreenItemData" at 68,78 size 158x20; Text 'HMI device type:'
   TextField "HmiScreenItemData_1" at 230,78 size 246x20; Text 'KTP400 Basic+ PN 15.1.0.0'
   TextField "HmiScreenItemData_2" at 68,99 size 158x20; Text 'Connection:'
   TextField "HmiScreenItemData_3" at 230,99 size 246x20; Text 'PROFINET (X1)'
   TextField "HmiScreenItemData_4" at 68,120 size 158x20; Text 'PLC:'
   TextField "HmiScreenItemData_5" at 230,120 size 246x20; Text 'SIMATIC S7 1200'
   Button "Back" at 65,46 size 136x30; TextOff 'Back'
      on Release: ActivateScreen("System screens", 0)
*)